// TIA Portal project "FK_PiPl" (V16) (continued)
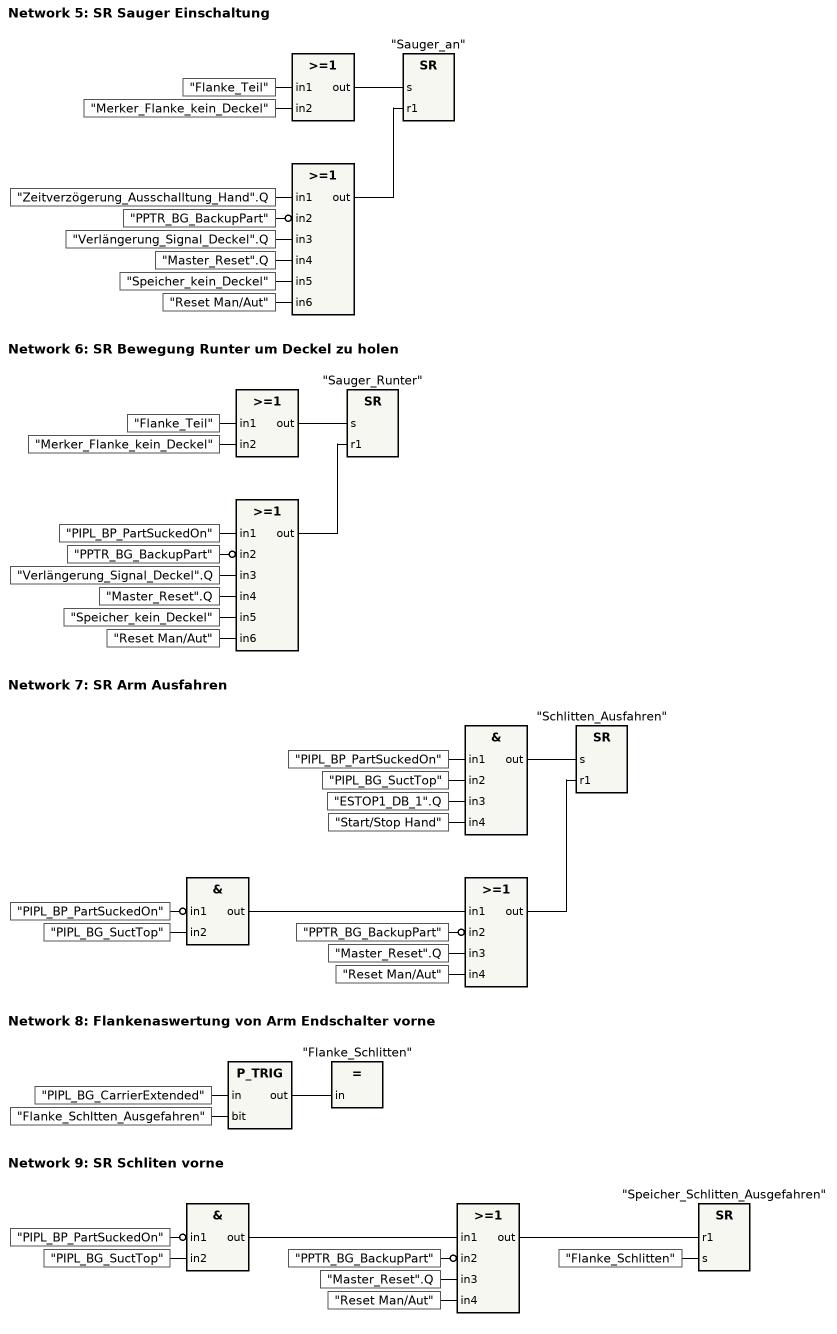
   IF "Flanke_Teil" OR "Merker_Flanke_kein_Deckel" THEN
       "Sauger_an" := TRUE;   // SR flip-flop
   END_IF;
   IF "Zeitverzögerung_Ausschalltung_Hand".Q OR NOT "PPTR_BG_BackupPart" OR "Verlängerung_Signal_Deckel".Q OR "Master_Reset".Q OR "Speicher_kein_Deckel" OR "Reset Man/Aut" THEN
       "Sauger_an" := FALSE;
   END_IF;
END_REGION

REGION Network 6: SR Bewegung Runter um Deckel zu holen
   IF "Flanke_Teil" OR "Merker_Flanke_kein_Deckel" THEN
       "Sauger_Runter" := TRUE;   // SR flip-flop
   END_IF;
   IF "PIPL_BP_PartSuckedOn" OR NOT "PPTR_BG_BackupPart" OR "Verlängerung_Signal_Deckel".Q OR "Master_Reset".Q OR "Speicher_kein_Deckel" OR "Reset Man/Aut" THEN
       "Sauger_Runter" := FALSE;
   END_IF;
END_REGION

REGION Network 7: SR Arm Ausfahren
   IF "PIPL_BP_PartSuckedOn" AND "PIPL_BG_SuctTop" AND "ESTOP1_DB_1".Q AND "Start/Stop Hand" THEN
       "Schlitten_Ausfahren" := TRUE;   // SR flip-flop
   END_IF;
   IF (NOT "PIPL_BP_PartSuckedOn" AND "PIPL_BG_SuctTop") OR NOT "PPTR_BG_BackupPart" OR "Master_Reset".Q OR "Reset Man/Aut" THEN
       "Schlitten_Ausfahren" := FALSE;
   END_IF;
END_REGION

REGION Network 8: Flankenaswertung von Arm Endschalter vorne
   #_w1 := "PIPL_BG_CarrierExtended" AND NOT "Flanke_Schltten_Ausgefahren";   // rising edge
   "Flanke_Schltten_Ausgefahren" := "PIPL_BG_CarrierExtended";
   "Flanke_Schlitten" := #_w1;
END_REGION

REGION Network 9: SR Schliten vorne
   IF "Flanke_Schlitten" THEN
       "Speicher_Schlitten_Ausgefahren" := TRUE;   // SR flip-flop
   END_IF;
   IF (NOT "PIPL_BP_PartSuckedOn" AND "PIPL_BG_SuctTop") OR NOT "PPTR_BG_BackupPart" OR "Master_Reset".Q OR "Reset Man/Aut" THEN
       "Speicher_Schlitten_Ausgefahren" := FALSE;
   END_IF;
END_REGION

REGION Network 10: Zeitverzögerung von Saugerabschaltung
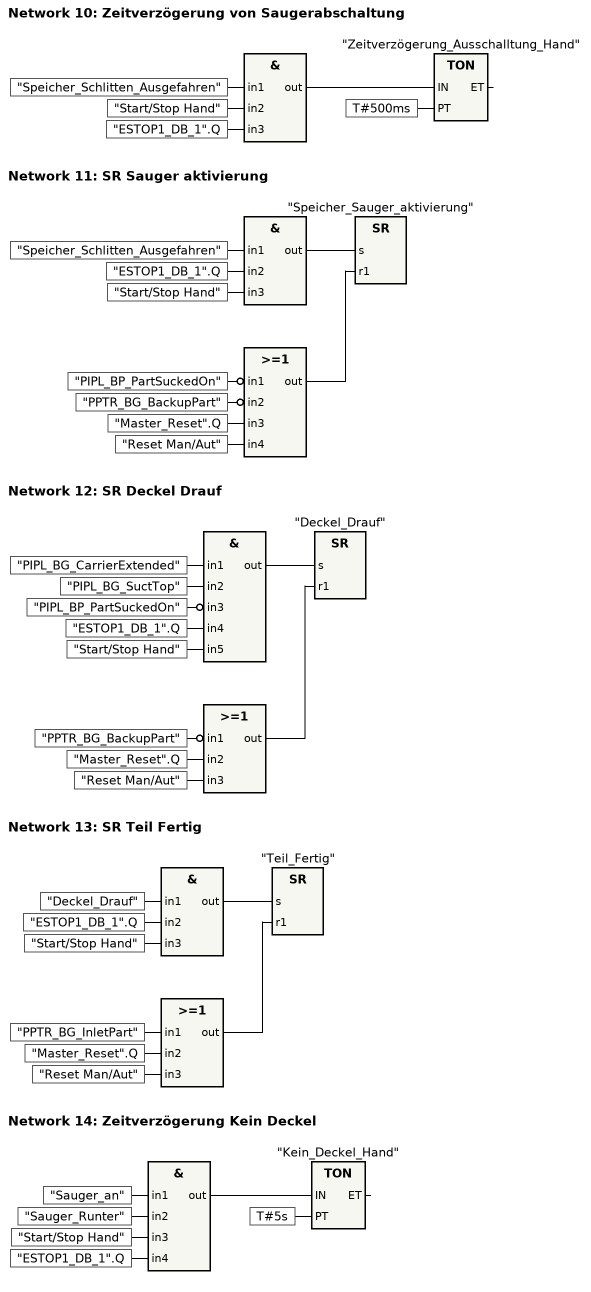
   "Zeitverzögerung_Ausschalltung_Hand".TON(IN := "Speicher_Schlitten_Ausgefahren" AND "Start/Stop Hand" AND "ESTOP1_DB_1".Q,
                           PT := T#500ms);
END_REGION

REGION Network 11: SR Sauger aktivierung
   IF "Speicher_Schlitten_Ausgefahren" AND "ESTOP1_DB_1".Q AND "Start/Stop Hand" THEN
       "Speicher_Sauger_aktivierung" := TRUE;   // SR flip-flop
   END_IF;
   IF NOT "PIPL_BP_PartSuckedOn" OR NOT "PPTR_BG_BackupPart" OR "Master_Reset".Q OR "Reset Man/Aut" THEN
       "Speicher_Sauger_aktivierung" := FALSE;
   END_IF;
END_REGION

REGION Network 12: SR Deckel Drauf
   IF "PIPL_BG_CarrierExtended" AND "PIPL_BG_SuctTop" AND NOT "PIPL_BP_PartSuckedOn" AND "ESTOP1_DB_1".Q AND "Start/Stop Hand" THEN
       "Deckel_Drauf" := TRUE;   // SR flip-flop
   END_IF;
   IF NOT "PPTR_BG_BackupPart" OR "Master_Reset".Q OR "Reset Man/Aut" THEN "Deckel_Drauf" := FALSE; END_IF;
END_REGION

REGION Network 13: SR Teil Fertig
   IF "Deckel_Drauf" AND "ESTOP1_DB_1".Q AND "Start/Stop Hand" THEN
       "Teil_Fertig" := TRUE;   // SR flip-flop
   END_IF;
   IF "PPTR_BG_InletPart" OR "Master_Reset".Q OR "Reset Man/Aut" THEN "Teil_Fertig" := FALSE; END_IF;
END_REGION

REGION Network 14: Zeitverzögerung Kein Deckel
   // Wenn nach der eingestellten Zeit kein Deckel angesaugt wurde gibt die Maschine ein Fehler aus
   "Kein_Deckel_Hand".TON(IN := "Sauger_an" AND "Sauger_Runter" AND "Start/Stop Hand" AND "ESTOP1_DB_1".Q,
                          PT := T#5s);
END_REGION

REGION Network 15: SR kein Deckel
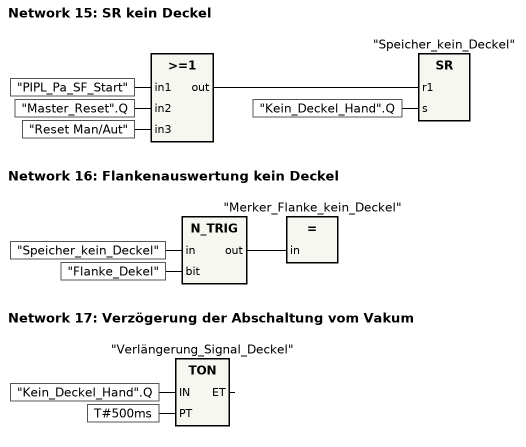
   IF "Kein_Deckel_Hand".Q THEN
       "Speicher_kein_Deckel" := TRUE;   // SR flip-flop
   END_IF;
   IF "PIPL_Pa_SF_Start" OR "Master_Reset".Q OR "Reset Man/Aut" THEN "Speicher_kein_Deckel" := FALSE; END_IF;
END_REGION

REGION Network 16: Flankenauswertung kein Deckel
   #_w1 := NOT "Speicher_kein_Deckel" AND "Flanke_Dekel";   // falling edge
   "Flanke_Dekel" := "Speicher_kein_Deckel";
   "Merker_Flanke_kein_Deckel" := #_w1;
END_REGION

REGION Network 17: Verzögerung der Abschaltung vom Vakum
   "Verlängerung_Signal_Deckel".TON(IN := "Kein_Deckel_Hand".Q, PT := T#500ms);
END_REGION
END_FUNCTION

FUNCTION "Druck" : Void   // FC6, FBD
{ S7_Optimized_Access := 'TRUE' }
VERSION : 0.1
BEGIN

REGION Network 1: Drucksensor Auslesung
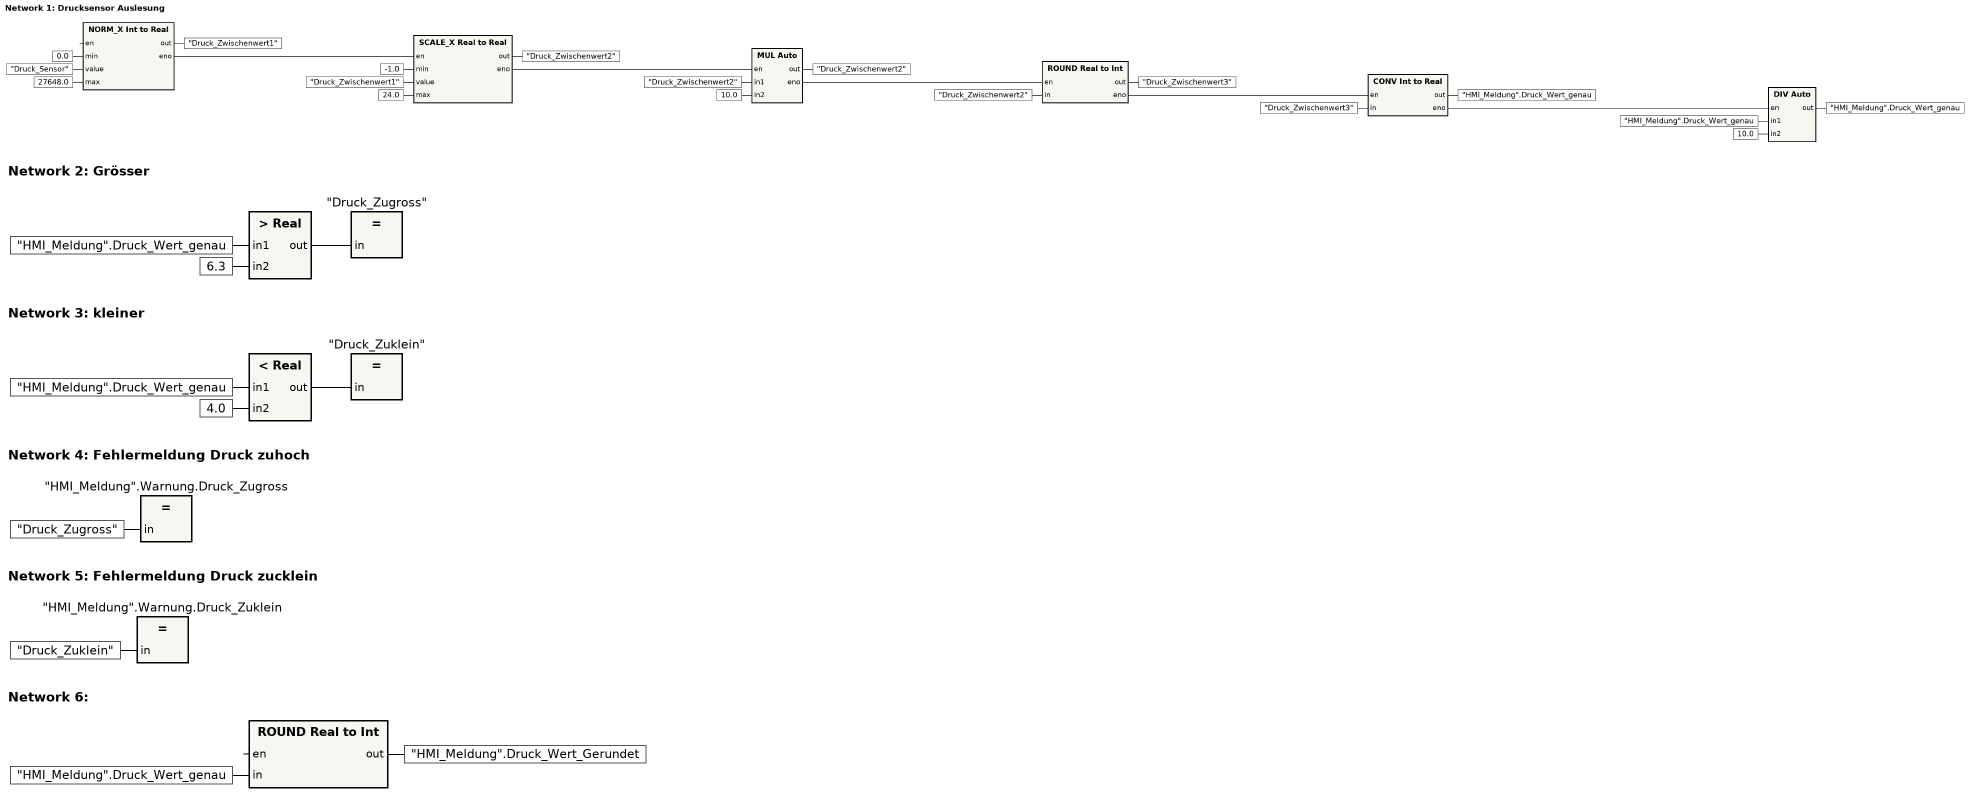
   "Druck_Zwischenwert1" := NORM_X(MIN := 0.0, VALUE := "Druck_Sensor", MAX := 27648.0);
   "Druck_Zwischenwert2" := SCALE_X(MIN := -1.0, VALUE := "Druck_Zwischenwert1", MAX := 24.0);
   "Druck_Zwischenwert2" := "Druck_Zwischenwert2" * 10.0;
   "Druck_Zwischenwert3" := ROUND("Druck_Zwischenwert2");
   "HMI_Meldung".Druck_Wert_genau := INT_TO_REAL("Druck_Zwischenwert3");
   "HMI_Meldung".Druck_Wert_genau := "HMI_Meldung".Druck_Wert_genau / 10.0;
END_REGION

REGION Network 2: Grösser
   "Druck_Zugross" := "HMI_Meldung".Druck_Wert_genau > 6.3;
END_REGION

REGION Network 3: kleiner
   "Druck_Zuklein" := "HMI_Meldung".Druck_Wert_genau < 4.0;
END_REGION

REGION Network 4: Fehlermeldung Druck zuhoch
   "HMI_Meldung".Warnung.Druck_Zugross := "Druck_Zugross";
END_REGION

REGION Network 5: Fehlermeldung Druck zucklein
   "HMI_Meldung".Warnung.Druck_Zuklein := "Druck_Zuklein";
END_REGION

REGION Network 6
   "HMI_Meldung".Druck_Wert_Gerundet := ROUND("HMI_Meldung".Druck_Wert_genau);
END_REGION
END_FUNCTION

FUNCTION "Ausgänge" : Void   // FC8, FBD
{ S7_Optimized_Access := 'TRUE' }
VERSION : 0.1
BEGIN

REGION Network 1: Pick&Placer Sauger nach unten (125MB3)
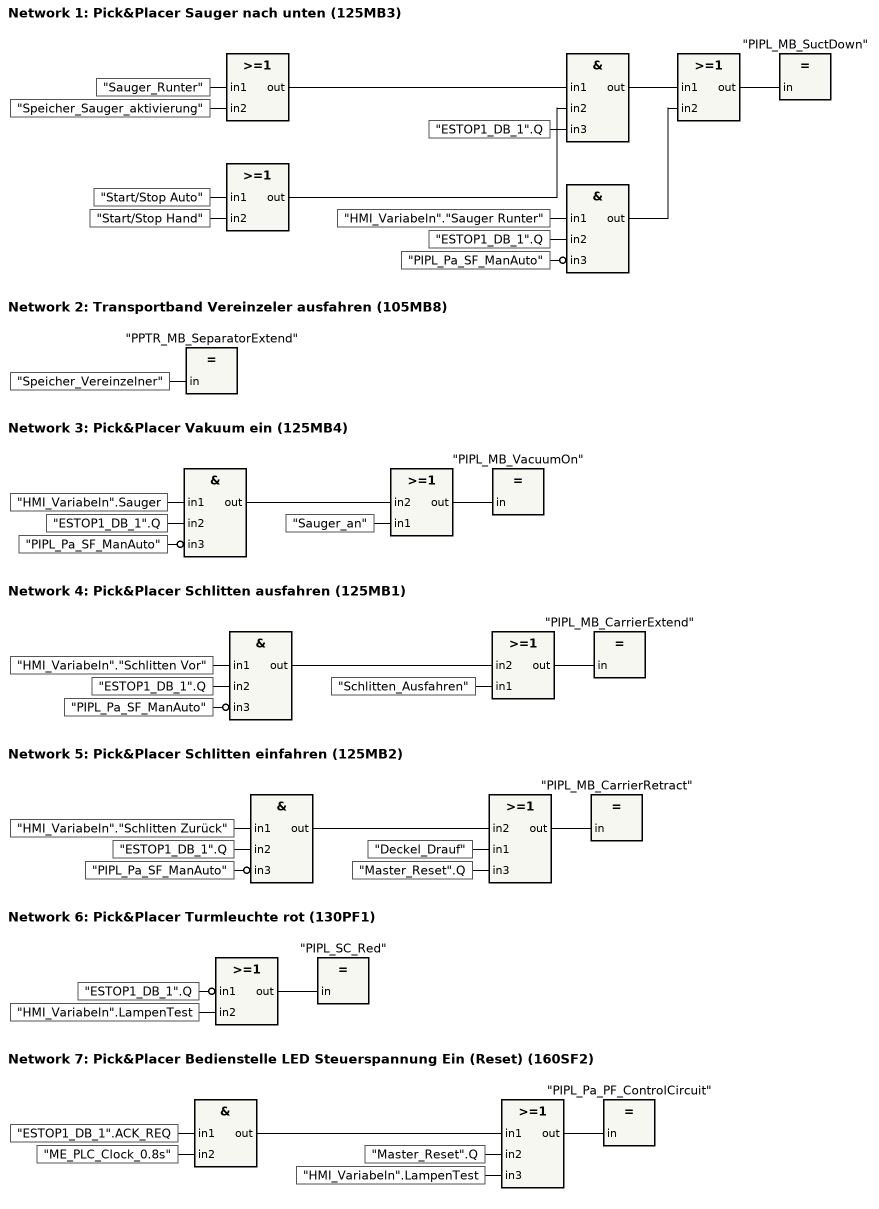
   "PIPL_MB_SuctDown" := (("Sauger_Runter" OR "Speicher_Sauger_aktivierung") AND ("Start/Stop Auto" OR "Start/Stop Hand") AND "ESTOP1_DB_1".Q) OR ("HMI_Variabeln"."Sauger Runter" AND "ESTOP1_DB_1".Q AND NOT "PIPL_Pa_SF_ManAuto");
END_REGION

REGION Network 2: Transportband Vereinzeler ausfahren (105MB8)
   "PPTR_MB_SeparatorExtend" := "Speicher_Vereinzelner";
END_REGION

REGION Network 3: Pick&Placer Vakuum ein (125MB4)
   "PIPL_MB_VacuumOn" := ("HMI_Variabeln".Sauger AND "ESTOP1_DB_1".Q AND NOT "PIPL_Pa_SF_ManAuto") OR "Sauger_an";
END_REGION

REGION Network 4: Pick&Placer Schlitten ausfahren (125MB1)
   "PIPL_MB_CarrierExtend" := ("HMI_Variabeln"."Schlitten Vor" AND "ESTOP1_DB_1".Q AND NOT "PIPL_Pa_SF_ManAuto") OR "Schlitten_Ausfahren";
END_REGION

REGION Network 5: Pick&Placer Schlitten einfahren (125MB2)
   "PIPL_MB_CarrierRetract" := ("HMI_Variabeln"."Schlitten Zurück" AND "ESTOP1_DB_1".Q AND NOT "PIPL_Pa_SF_ManAuto") OR "Deckel_Drauf" OR "Master_Reset".Q;
END_REGION

REGION Network 6: Pick&Placer Turmleuchte rot (130PF1)
   "PIPL_SC_Red" := NOT "ESTOP1_DB_1".Q OR "HMI_Variabeln".LampenTest;
END_REGION

REGION Network 7: Pick&Placer Bedienstelle LED Steuerspannung Ein (Reset) (160SF2)
   "PIPL_Pa_PF_ControlCircuit" := ("ESTOP1_DB_1".ACK_REQ AND "ME_PLC_Clock_0.8s") OR "Master_Reset".Q OR "HMI_Variabeln".LampenTest;
END_REGION

REGION Network 8: Pick&Placer Turmleuchte grün (130PF1)
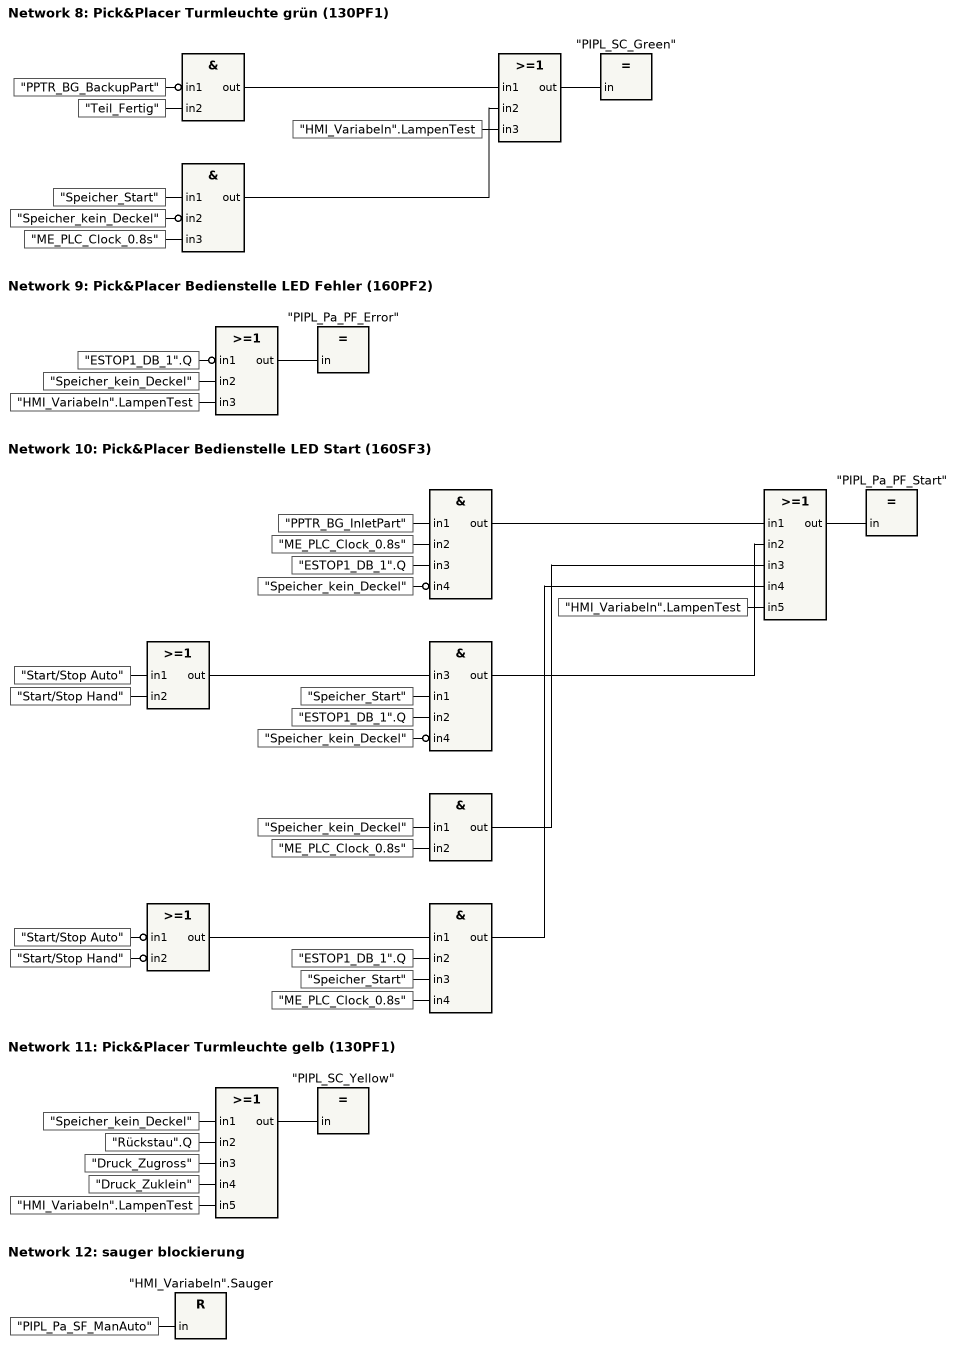
   "PIPL_SC_Green" := (NOT "PPTR_BG_BackupPart" AND "Teil_Fertig") OR ("Speicher_Start" AND NOT "Speicher_kein_Deckel" AND "ME_PLC_Clock_0.8s") OR "HMI_Variabeln".LampenTest;
END_REGION

REGION Network 9: Pick&Placer Bedienstelle LED Fehler (160PF2)
   "PIPL_Pa_PF_Error" := NOT "ESTOP1_DB_1".Q OR "Speicher_kein_Deckel" OR "HMI_Variabeln".LampenTest;
END_REGION

REGION Network 10: Pick&Placer Bedienstelle LED Start (160SF3)
   "PIPL_Pa_PF_Start" := ("PPTR_BG_InletPart" AND "ME_PLC_Clock_0.8s" AND "ESTOP1_DB_1".Q AND NOT "Speicher_kein_Deckel") OR (("Start/Stop Auto" OR "Start/Stop Hand") AND "Speicher_Start" AND "ESTOP1_DB_1".Q AND NOT "Speicher_kein_Deckel") OR ("Speicher_kein_Deckel" AND "ME_PLC_Clock_0.8s") OR ((NOT "Start/Stop Auto" OR NOT "Start/Stop Hand") AND "ESTOP1_DB_1".Q AND "Speicher_Start" AND "ME_PLC_Clock_0.8s") OR "HMI_Variabeln".LampenTest;
END_REGION

REGION Network 11: Pick&Placer Turmleuchte gelb (130PF1)
   "PIPL_SC_Yellow" := "Speicher_kein_Deckel" OR "Rückstau".Q OR "Druck_Zugross" OR "Druck_Zuklein" OR "HMI_Variabeln".LampenTest;
END_REGION

REGION Network 12: sauger blockierung
   IF "PIPL_Pa_SF_ManAuto" THEN "HMI_Variabeln".Sauger := FALSE; END_IF;
END_REGION

REGION Network 13: Vakurunter Blockierung
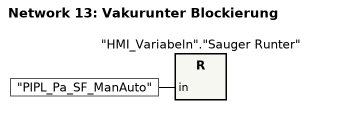
   IF "PIPL_Pa_SF_ManAuto" THEN "HMI_Variabeln"."Sauger Runter" := FALSE; END_IF;
END_REGION
END_FUNCTION

ORGANIZATION_BLOCK "Main"   // OB1, FBD, ProgramCycle
TITLE = "Main Program Sweep (Cycle)"
{ S7_Optimized_Access := 'TRUE' }
VERSION : 0.1
   VAR_INPUT
      Initial_Call : Bool;   // Initial call of this OB
      Remanence : Bool;   // =True, if remanent data are available
   END_VAR
BEGIN

REGION Network 1: initialisierung Ausgaenge
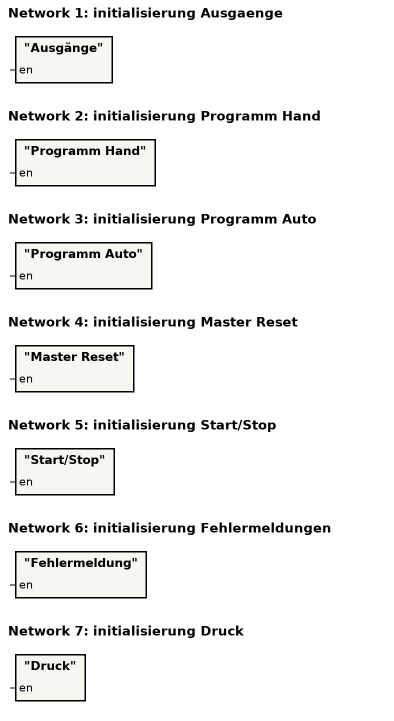
   "Ausgänge"();
END_REGION

REGION Network 2: initialisierung Programm Hand
   "Programm Hand"();
END_REGION

REGION Network 3: initialisierung Programm Auto
   "Programm Auto"();
END_REGION

REGION Network 4: initialisierung Master Reset
   "Master Reset"();
END_REGION

REGION Network 5: initialisierung Start/Stop
   "Start/Stop"();
END_REGION

REGION Network 6: initialisierung Fehlermeldungen
   "Fehlermeldung"();
END_REGION

REGION Network 7: initialisierung Druck
   "Druck"();
END_REGION
END_ORGANIZATION_BLOCK

(* ===== HMI "HMI_RT_1" =====
system functions are stored by id; their names below are inferred from use
connection "HMI_1": ETHERNET, S7_1500_OMS

HMI tags "Standard-Variablentabelle"
   "Variable_Bildnummer" : UInt, internal
   "Speicher_Start" : Bool = PLC Speicher_Start AT %M4.0, 1 s
   "HMI_Variabeln_Förderband vor" : Bool = PLC HMI_Variabeln."Förderband vor", 1 s
   "HMI_Variabeln_Förderbad Zurück" : Bool = PLC HMI_Variabeln."Förderbad Zurück", 1 s
   "HMI_Variabeln_Stop" : Bool = PLC HMI_Variabeln."Schlitten Vor", 1 s
   "HMI_Variabeln_Schlitten Zurück" : Bool = PLC HMI_Variabeln."Schlitten Zurück", 1 s
   "HMI_Variabeln_Sauger" : Bool = PLC HMI_Variabeln.Sauger, 1 s
   "HMI_Variabeln_Sauger Runter" : Bool = PLC HMI_Variabeln."Sauger Runter", 1 s
   "HMI_Variabeln_LampenTest" : Bool = PLC HMI_Variabeln.LampenTest, 1 s
   "HMI_Meldung_Druck_Wert_genau" : Real = PLC HMI_Meldung.Druck_Wert_genau AT %DB8.DBD2, 1 s

HMI tags "DB122"
   "Datenbaustein_1_Sammelstoerung" : Bool = PLC Datenbaustein_1.Sammelstoerung, 1 s
   "Datenbaustein_1_Lampe_Ein" : Bool = PLC Datenbaustein_1.Lampe_Ein, 1 s
   "Datenbaustein_1_Lampe_Aus" : Bool = PLC Datenbaustein_1.Lampe_Aus, 1 s
   "Datenbaustein_1_Reserve3" : Bool = PLC Datenbaustein_1.Reserve3, 1 s
   "Datenbaustein_1_Reserve4" : Bool = PLC Datenbaustein_1.Reserve4, 1 s
   "Datenbaustein_1_Reserve5" : Bool = PLC Datenbaustein_1.Reserve5, 1 s
   "Datenbaustein_1_Reserve6" : Bool = PLC Datenbaustein_1.Reserve6, 1 s
   "Datenbaustein_1_Reserve7" : Bool = PLC Datenbaustein_1.Reserve7, 1 s
   "Datenbaustein_1_Reserve8" : Bool = PLC Datenbaustein_1.Reserve8, 1 s
   "Datenbaustein_1_Reserve9" : Bool = PLC Datenbaustein_1.Reserve9, 1 s
   "Datenbaustein_1_Wert" : Int = PLC Datenbaustein_1.Wert, 1 s

HMI tags "Meldung"
   "Fehler" : Int AT %DB8.DBW8, 1 s
   "Warnung" : Int AT %DB8.DBW6, 1 s
   "Meldungen" : Int AT %DB8.DBW10, 1 s
   "Druck_Wert_Genau" : Real AT %DB8.DBD2, 1 s
   "Druck_Wert_gerundet" : Int AT %DB8.DBW0, 1 s

discrete alarms
   1: 'Kein Deckel vorhanden', class Errors, trigger "Fehler" bit 8
   2: 'Not-Aus betätigt', class Errors, trigger "Fehler" bit 9
   3: 'Not-Aus Quitieren', class Errors, trigger "Warnung" bit 8
   4: 'Werkstück erkannt/bereit', class Errors, trigger "Meldungen" bit 8
   5: 'Rückstau zu gross', class Errors, trigger "Warnung" bit 9
   6: 'Druck zuhoch', class Errors, trigger "Warnung" bit 10
   7: 'Druck zuklein', class Errors, trigger "Warnung" bit 11

text list "Textliste_Bildnamen": 1 'Grundbild'

screen "Home" 480x272
   Button "Schaltfläche_1" at 384,232 size 96x40; TextOff 'Text'; PictureOff "Right_Arrow"
      on Press: ActivateScreen("Pamasol_Info", 0)
   Button "Schaltfläche_4" at 0,232 size 96x40; TextOff 'Text'; PictureOff "Left_Arrow"
      on Press: ActivateScreen("Manuelle_Bedienung", 0)
   Button "Schaltfläche_2" at 8,0 size 304x80; TextOff 'Text'; PictureOff "PWMA_Logo"
   GraphicView "Grafikanzeige_1" at 270,-1 size 208x80; Picture "bg-top-3104a5681f3727e8357f577a4a6a55f0"
   Clock "Uhr_1" at 104,88 size 120x120
   Gauge "Zeigerinstrument_1" at 264,88 size 120x120; CaptionText 'Druck'; UnitText 'Bar'
      ProcessValue <- "Druck_Wert_Genau"
   IOField "EA-Feld_1" at 202,233 size 73x39; FormatPattern 99.9
      ProcessValue <- "HMI_Meldung_Druck_Wert_genau"
      Visibility <- "Druck_Wert_gerundet"
   Button "Schaltfläche_19" at 239,238 size 33x29; TextOff 'Bar'

screen "Pamasol_Info" 480x272
   Button "Schaltfläche_1" at 24,80 size 168x24; TextOff 'Pamasol Willi Mäder AG'
   Button "Schaltfläche_2" at 24,104 size 168x24; TextOff 'Driesbülstr.2'
   Button "Schaltfläche_3" at 24,128 size 168x24; TextOff '8808 Pfäffikon / SZ'
   Button "Schaltfläche_4" at 24,152 size 168x24; TextOff 'CH-Swizerland'
   Button "Schaltfläche_5" at 224,80 size 64x24; TextOff 'Tel.:'
   Button "Schaltfläche_6" at 224,104 size 64x24; TextOff 'Fax:'
   Button "Schaltfläche_7" at 224,128 size 64x24; TextOff 'E-mail:'
   Button "Schaltfläche_8" at 224,152 size 80x24; TextOff 'Hompage:'
   Button "Schaltfläche_9" at 328,80 size 128x24; TextOff '+41 55 417 40 40'
   Button "Schaltfläche_10" at 328,104 size 128x24; TextOff '+41 55 417 40 44'
   Button "Schaltfläche_11" at 328,128 size 128x24; TextOff 'info@pamasol.com'
   Button "Schaltfläche_12" at 328,152 size 128x24; TextOff 'www.pamasol.com'
   GraphicView "Grafikanzeige_2" at 256,0 size 198x68; Picture "bg-top-3104a5681f3727e8357f577a4a6a55f0"
   GraphicView "Grafikanzeige_1" at 40,0 size 224x64; Picture "PWMA_Logo"
   Button "Schaltfläche_13" at 24,192 size 64x16; TextOff 'Machines:'
   Button "Schaltfläche_14" at 24,208 size 64x16; TextOff 'Date:'
   Button "Schaltfläche_15" at 256,192 size 128x16; TextOff 'Pick and Placer-Modul'
   Button "Schaltfläche_16" at 256,208 size 128x16; TextOff '13.07.22'
   Button "Schaltfläche_17" at 384,232 size 96x40; TextOff 'Text'; PictureOff "Right_Arrow"
      on Press: ActivateScreen("Meldungen", 0)
   Button "Schaltfläche_18" at 0,232 size 96x40; TextOff 'Text'; PictureOff "Left_Arrow"
      on Press: ActivateScreen("Home", 0)
   IOField "EA-Feld_1" at 202,233 size 73x39; FormatPattern 99.9
      ProcessValue <- "HMI_Meldung_Druck_Wert_genau"
      Visibility <- "Druck_Wert_gerundet"
   Button "Schaltfläche_19" at 239,238 size 33x29; TextOff 'Bar'

screen "Meldungen" 480x272
   AlarmView "Meldeanzeige_1" at 0,8 size 480x224
   Button "Schaltfläche_17" at 384,232 size 96x40; TextOff 'Text'; PictureOff "Right_Arrow"
      on Press: ActivateScreen("Manuelle_Bedienung", 0)
   Button "Schaltfläche_18" at 0,232 size 96x40; TextOff 'Text'; PictureOff "Left_Arrow"
      on Press: ActivateScreen("Pamasol_Info", 0)
   IOField "EA-Feld_1" at 202,233 size 73x39; FormatPattern 99.9
      Visibility <- "Druck_Wert_gerundet"
      ProcessValue <- "HMI_Meldung_Druck_Wert_genau"
   Button "Schaltfläche_19" at 239,238 size 33x29; TextOff 'Bar'

screen "Manuelle_Bedienung" 480x272
   Button "Schaltfläche_1" at 40,32 size 104x32; TextOff 'Transportband'
   Button "Schaltfläche_2" at 16,72 size 64x32; TextOff 'Vor'
      on Press: SetBit("HMI_Variabeln_Förderband vor")
      on Release: ResetBit("HMI_Variabeln_Förderband vor")
   Button "Schaltfläche_3" at 96,72 size 64x32; TextOff 'Zurück'
      on Press: SetBit("HMI_Variabeln_Förderbad Zurück")
      on Release: ResetBit("HMI_Variabeln_Förderbad Zurück")
   Button "Schaltfläche_4" at 384,232 size 96x40; TextOff 'Text'; PictureOff "Right_Arrow"
      on Press: ActivateScreen("Home", 0); ResetBit("HMI_Variabeln_LampenTest"); ResetBit("HMI_Variabeln_Förderband vor"); ResetBit("HMI_Variabeln_Förderbad Zurück"); ResetBit("HMI_Variabeln_Stop"); SetBit("HMI_Variabeln_Schlitten Zurück"); ResetBit("HMI_Variabeln_Sauger"); ResetBit("HMI_Variabeln_Sauger Runter")
   Button "Schaltfläche_5" at 0,232 size 96x40; TextOff 'Text'; PictureOff "Left_Arrow"
      on Press: ActivateScreen("Meldungen", 0); ResetBit("HMI_Variabeln_LampenTest"); ResetBit("HMI_Variabeln_Förderband vor"); ResetBit("HMI_Variabeln_Förderbad Zurück"); ResetBit("HMI_Variabeln_Sauger"); ResetBit("HMI_Variabeln_Stop"); SetBit("HMI_Variabeln_Schlitten Zurück"); ResetBit("HMI_Variabeln_Sauger Runter")
   Button "Schaltfläche_6" at 176,8 size 152x32; TextOff 'Manuelle Ansteuerung'
   Button "Schaltfläche_7" at 344,32 size 104x32; TextOff 'Schlitten'
   Button "Schaltfläche_8" at 320,72 size 64x32; TextOff 'Vor'
      on Release: ResetBit("HMI_Variabeln_Stop")
      on Press: SetBit("HMI_Variabeln_Stop"); ResetBit("HMI_Variabeln_Schlitten Zurück")
   Button "Schaltfläche_9" at 400,72 size 64x32; TextOff 'Zurück'
      on Release: ResetBit("HMI_Variabeln_Schlitten Zurück")
      on Press: SetBit("HMI_Variabeln_Schlitten Zurück"); ResetBit("HMI_Variabeln_Stop")
   Button "Schaltfläche_10" at 40,136 size 104x32; TextOff 'Vakum'
   Button "Schaltfläche_11" at 16,176 size 64x32; TextOff 'An'
      on Press: SetBit("HMI_Variabeln_Sauger")
   Button "Schaltfläche_12" at 104,176 size 64x32; TextOff 'Aus'
      on Press: ResetBit("HMI_Variabeln_Sauger")
   Button "Schaltfläche_13" at 344,136 size 104x32; TextOff 'Vakum'
   Button "Schaltfläche_14" at 320,176 size 64x32; TextOff 'Hoch'
      on Press: ResetBit("HMI_Variabeln_Sauger Runter")
   Button "Schaltfläche_15" at 408,176 size 64x32; TextOff 'Runter'
      on Press: SetBit("HMI_Variabeln_Sauger Runter")
   Button "Schaltfläche_16" at 193,77 size 96x32; TextOff 'Lampentest'
   Button "Schaltfläche_17" at 208,123 size 64x32; TextOff 'An'
      on Press: SetBit("HMI_Variabeln_LampenTest")
      on Release: ResetBit("HMI_Variabeln_LampenTest")
   IOField "EA-Feld_1" at 202,233 size 73x39; FormatPattern 99.9
      ProcessValue <- "HMI_Meldung_Druck_Wert_genau"
      Visibility <- "Druck_Wert_gerundet"
   Button "Schaltfläche_19" at 239,238 size 33x29; TextOff 'Bar'
*)